// TIA Portal project "OP-TQ-01" (V13) (continued)
REGION Network 24: RESET ALARME DE SINAL ANALÓGICO
   RUNG wire#powerrail
      I_Contact( #Alarms.LL )
      I_Contact( #Alarms.L )
      I_Contact( #Alarms.H )
      I_Contact( #Alarms.HH )
      Contact( #RESET )
      wire#w1
      R_Coil( #AnalogInputAlarm )
   END_RUNG
   RUNG wire#powerrail
      Contact( #UnableAlarms )
   END_RUNG wire#w1
   RUNG wire#powerrail
      Contact( #Maint )
   END_RUNG wire#w1
   // the same network as SCL:
   IF (NOT #Alarms.LL AND NOT #Alarms.L AND NOT #Alarms.H AND NOT #Alarms.HH AND #RESET) OR #UnableAlarms OR #Maint THEN
       #AnalogInputAlarm := FALSE;
   END_IF;
END_REGION

REGION Network 25: 0 - STATUS OK
   RUNG wire#powerrail
      I_Contact( #AnalogInputFault )
      I_Contact( #AnalogInputAlarm )
      Contact( #Maint )
      { S7_GenerateENO := "TRUE" } Move(in := 0, out1 => #Status)
   END_RUNG
   // the same network as SCL:
   IF NOT #AnalogInputFault AND NOT #AnalogInputAlarm AND #Maint THEN #Status := 0; END_IF;
END_REGION

REGION Network 26: 1 - STATUS FALHA - UNDER FLOW
   RUNG wire#powerrail
      Contact( #Alarms.UDF )
      Contact( #Maint )
      { S7_GenerateENO := "TRUE" } Move(in := 1, out1 => #Status)
   END_RUNG
   // the same network as SCL:
   IF #Alarms.UDF AND #Maint THEN #Status := 1; END_IF;
END_REGION

REGION Network 27: 2 - STATUS FALHA - UNDER RANGE
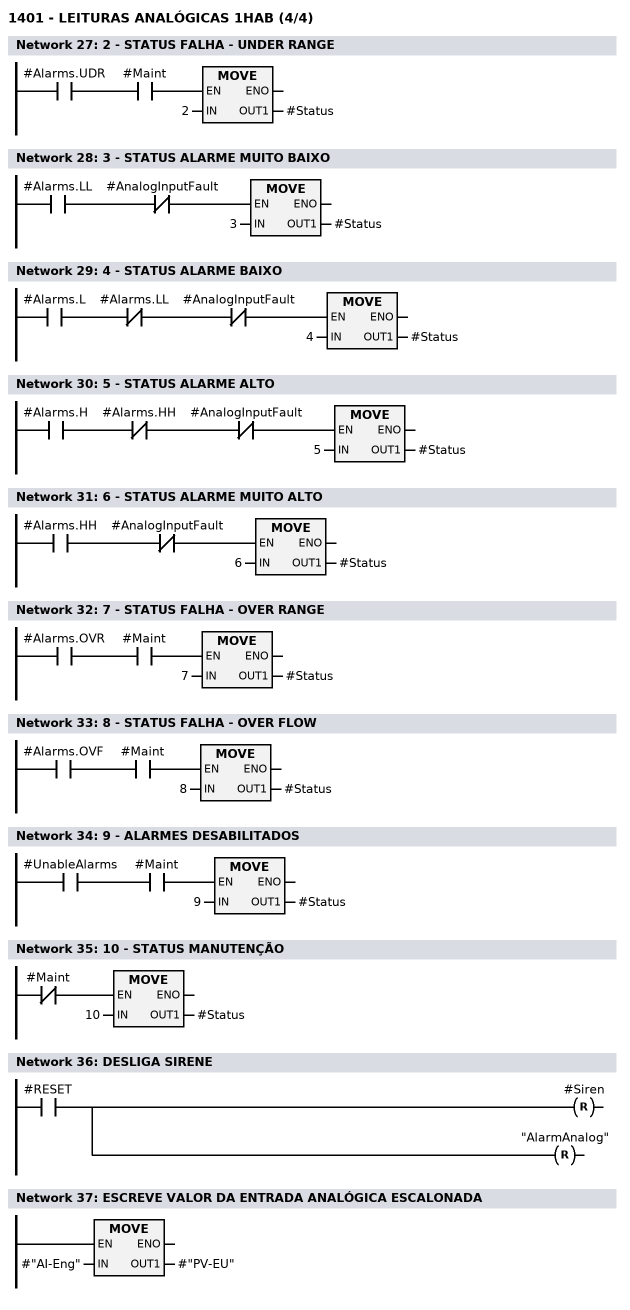
   RUNG wire#powerrail
      Contact( #Alarms.UDR )
      Contact( #Maint )
      { S7_GenerateENO := "TRUE" } Move(in := 2, out1 => #Status)
   END_RUNG
   // the same network as SCL:
   IF #Alarms.UDR AND #Maint THEN #Status := 2; END_IF;
END_REGION

REGION Network 28: 3 - STATUS ALARME MUITO BAIXO
   RUNG wire#powerrail
      Contact( #Alarms.LL )
      I_Contact( #AnalogInputFault )
      { S7_GenerateENO := "TRUE" } Move(in := 3, out1 => #Status)
   END_RUNG
   // the same network as SCL:
   IF #Alarms.LL AND NOT #AnalogInputFault THEN #Status := 3; END_IF;
END_REGION

REGION Network 29: 4 - STATUS ALARME BAIXO
   RUNG wire#powerrail
      Contact( #Alarms.L )
      I_Contact( #Alarms.LL )
      I_Contact( #AnalogInputFault )
      { S7_GenerateENO := "TRUE" } Move(in := 4, out1 => #Status)
   END_RUNG
   // the same network as SCL:
   IF #Alarms.L AND NOT #Alarms.LL AND NOT #AnalogInputFault THEN #Status := 4; END_IF;
END_REGION

REGION Network 30: 5 - STATUS ALARME ALTO
   RUNG wire#powerrail
      Contact( #Alarms.H )
      I_Contact( #Alarms.HH )
      I_Contact( #AnalogInputFault )
      { S7_GenerateENO := "TRUE" } Move(in := 5, out1 => #Status)
   END_RUNG
   // the same network as SCL:
   IF #Alarms.H AND NOT #Alarms.HH AND NOT #AnalogInputFault THEN #Status := 5; END_IF;
END_REGION

REGION Network 31: 6 - STATUS ALARME MUITO ALTO
   RUNG wire#powerrail
      Contact( #Alarms.HH )
      I_Contact( #AnalogInputFault )
      { S7_GenerateENO := "TRUE" } Move(in := 6, out1 => #Status)
   END_RUNG
   // the same network as SCL:
   IF #Alarms.HH AND NOT #AnalogInputFault THEN #Status := 6; END_IF;
END_REGION

REGION Network 32: 7 - STATUS FALHA - OVER RANGE
   RUNG wire#powerrail
      Contact( #Alarms.OVR )
      Contact( #Maint )
      { S7_GenerateENO := "TRUE" } Move(in := 7, out1 => #Status)
   END_RUNG
   // the same network as SCL:
   IF #Alarms.OVR AND #Maint THEN #Status := 7; END_IF;
END_REGION

REGION Network 33: 8 - STATUS FALHA - OVER FLOW
   RUNG wire#powerrail
      Contact( #Alarms.OVF )
      Contact( #Maint )
      { S7_GenerateENO := "TRUE" } Move(in := 8, out1 => #Status)
   END_RUNG
   // the same network as SCL:
   IF #Alarms.OVF AND #Maint THEN #Status := 8; END_IF;
END_REGION

REGION Network 34: 9 - ALARMES DESABILITADOS
   RUNG wire#powerrail
      Contact( #UnableAlarms )
      Contact( #Maint )
      { S7_GenerateENO := "TRUE" } Move(in := 9, out1 => #Status)
   END_RUNG
   // the same network as SCL:
   IF #UnableAlarms AND #Maint THEN #Status := 9; END_IF;
END_REGION

REGION Network 35: 10 - STATUS MANUTENÇÃO
   RUNG wire#powerrail
      I_Contact( #Maint )
      { S7_GenerateENO := "TRUE" } Move(in := 10, out1 => #Status)
   END_RUNG
   // the same network as SCL:
   IF NOT #Maint THEN #Status := 10; END_IF;
END_REGION

REGION Network 36: DESLIGA SIRENE
   RUNG wire#powerrail
      Contact( #RESET )
      wire#w1
      R_Coil( #Siren )
   END_RUNG
   RUNG wire#w1
      R_Coil( "AlarmAnalog" )
   END_RUNG
   // the same network as SCL:
   IF #RESET THEN
       #Siren := FALSE;
       "AlarmAnalog" := FALSE;
   END_IF;
END_REGION

REGION Network 37: ESCREVE VALOR DA ENTRADA ANALÓGICA ESCALONADA
   RUNG wire#powerrail
      { S7_GenerateENO := "TRUE" } Move(in := #"AI-Eng", out1 => #"PV-EU")
   END_RUNG
   // the same network as SCL:
   #"PV-EU" := #"AI-Eng";
END_REGION
END_FUNCTION_BLOCK

FUNCTION "1500 - SP-TT" : Void   // FC1500, LAD
{ S7_Optimized_Access := 'FALSE' }
VERSION : 0.1
   VAR_TEMP   // added for the SCL form of the ladder/FBD networks
      _w1 : Bool;
   END_VAR
BEGIN

REGION Network 1: VERIFICA TEMPERATURA MAX MAIOR QUE MIN
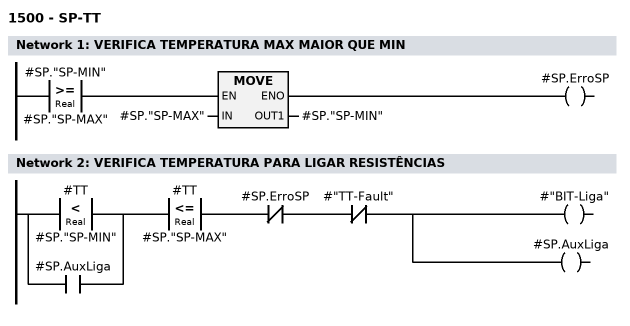
   RUNG wire#powerrail
      { S7_Templates := "SrcType := Real" } GE_Contact(in1 := #SP."SP-MIN", in2 := #SP."SP-MAX")
      { S7_GenerateENO := "TRUE" } Move(in := #SP."SP-MAX", out1 => #SP."SP-MIN")
      Coil( #SP.ErroSP )
   END_RUNG
   // the same network as SCL:
   // ENO of a box is taken as its EN; it also drops when the box reports an error
   #_w1 := #SP."SP-MIN" >= #SP."SP-MAX";
   IF #_w1 THEN #SP."SP-MIN" := #SP."SP-MAX"; END_IF;
   #SP.ErroSP := #_w1;
END_REGION

REGION Network 2: VERIFICA TEMPERATURA PARA LIGAR RESISTÊNCIAS
   RUNG wire#powerrail
      { S7_Templates := "SrcType := Real" } LT_Contact(in1 := #TT, in2 := #SP."SP-MIN")
      wire#w1
      { S7_Templates := "SrcType := Real" } LE_Contact(in1 := #TT, in2 := #SP."SP-MAX")
      I_Contact( #SP.ErroSP )
      I_Contact( #"TT-Fault" )
      wire#w2
      Coil( #"BIT-Liga" )
   END_RUNG
   RUNG wire#powerrail
      Contact( #SP.AuxLiga )
   END_RUNG wire#w1
   RUNG wire#w2
      Coil( #SP.AuxLiga )
   END_RUNG
   // the same network as SCL:
   #"BIT-Liga" := ((#TT < #SP."SP-MIN") OR #SP.AuxLiga) AND (#TT <= #SP."SP-MAX") AND NOT #SP.ErroSP AND NOT #"TT-Fault";
   #SP.AuxLiga := #"BIT-Liga";
END_REGION
END_FUNCTION

(* ===== HMI "HMI_RT_1" =====
connection "HMI_Connection_1": ETHERNET, S7_1200_OMS

HMI tags "Default tag table"
   "REC_ALM" : Bool = PLC "REC_ALM", 1 s
   "TT-006-R01A_AlarmsSts" : Alm-Bits, 1 s
   "TT-007-R01B_AlarmsSts" : Alm-Bits, 1 s
   "TT-008-R01C_AlarmsSts" : Alm-Bits, 1 s
   "TT-009-R01D_AlarmsSts" : Alm-Bits, 1 s
   "TT-010-R01E_AlarmsSts" : Alm-Bits, 1 s
   "TT-011-R01F_AlarmsSts" : Alm-Bits, 1 s
   "LT-009_AlarmsSts" : Alm-Bits, 1 s
   "LT-008_AlarmsSts" : Alm-Bits, 1 s

HMI tags "TT-006-R01A"
   "TT-006-R01A_UnableAlarms" : Bool, 1 s
   "TT-006-R01A_EngMax" : Real, 1 s
   "TT-006-R01A_EngMin" : Real, 1 s
   "TT-006-R01A_SP-HH" : Real, 1 s
   "TT-006-R01A_SP-H" : Real, 1 s
   "TT-006-R01A_SP-L" : Real, 1 s
   "TT-006-R01A_SP-LL" : Real, 1 s
   "TT-006-R01A_DelayHH" : Time, 1 s
   "TT-006-R01A_DelayH" : Time, 1 s
   "TT-006-R01A_DelayL" : Time, 1 s
   "TT-006-R01A_DelayLL" : Time, 1 s
   "TT-006-R01A_Siren" : Bool, 1 s
   "TT-006-R01A_SupRESET" : Bool, 1 s
   "TT-006-R01A_maint" : Bool, 1 s
   "TT-006-R01A_AlarmsEnable" : Alm-Bits, 1 s
   "TT-006-R01A_Alarms" : Alm-Bits, 1 s
   "TT-006-R01A_AI-Eng" : Real, 1 s
   "TT-006-R01A_Status" : Int, 1 s
   "TT-006-R01A_AnalogInput" : Int, 1 s

HMI tags "TT-007-R01B"
   "TT-007-R01B_UnableAlarms" : Bool, 1 s
   "TT-007-R01B_EngMax" : Real, 1 s
   "TT-007-R01B_EngMin" : Real, 1 s
   "TT-007-R01B_SP-HH" : Real, 1 s
   "TT-007-R01B_SP-H" : Real, 1 s
   "TT-007-R01B_SP-L" : Real, 1 s
   "TT-007-R01B_SP-LL" : Real, 1 s
   "TT-007-R01B_DelayHH" : Time, 1 s
   "TT-007-R01B_DelayH" : Time, 1 s
   "TT-007-R01B_DelayL" : Time, 1 s
   "TT-007-R01B_DelayLL" : Time, 1 s
   "TT-007-R01B_Siren" : Bool, 1 s
   "TT-007-R01B_SupRESET" : Bool, 1 s
   "TT-007-R01B_maint" : Bool, 1 s
   "TT-007-R01B_AlarmsEnable" : Alm-Bits, 1 s
   "TT-007-R01B_Alarms" : Alm-Bits, 1 s
   "TT-007-R01B_AI-Eng" : Real, 1 s
   "TT-007-R01B_Status" : Int, 1 s
   "TT-007-R01B_AnalogInput" : Int, 1 s

HMI tags "TT-008-R01C"
   "TT-008-R01C_UnableAlarms" : Bool, 1 s
   "TT-008-R01C_EngMax" : Real, 1 s
   "TT-008-R01C_EngMin" : Real, 1 s
   "TT-008-R01C_SP-HH" : Real, 1 s
   "TT-008-R01C_SP-H" : Real, 1 s
   "TT-008-R01C_SP-L" : Real, 1 s
   "TT-008-R01C_SP-LL" : Real, 1 s
   "TT-008-R01C_DelayHH" : Time, 1 s
   "TT-008-R01C_DelayH" : Time, 1 s
   "TT-008-R01C_DelayL" : Time, 1 s
   "TT-008-R01C_DelayLL" : Time, 1 s
   "TT-008-R01C_Siren" : Bool, 1 s
   "TT-008-R01C_SupRESET" : Bool, 1 s
   "TT-008-R01C_maint" : Bool, 1 s
   "TT-008-R01C_AlarmsEnable" : Alm-Bits, 1 s
   "TT-008-R01C_Alarms" : Alm-Bits, 1 s
   "TT-008-R01C_AI-Eng" : Real, 1 s
   "TT-008-R01C_Status" : Int, 1 s
   "TT-008-R01C_AnalogInput" : Int, 1 s

HMI tags "TT-009-R01D"
   "TT-009-R01D_UnableAlarms" : Bool, 1 s
   "TT-009-R01D_EngMax" : Real, 1 s
   "TT-009-R01D_EngMin" : Real, 1 s
   "TT-009-R01D_SP-HH" : Real, 1 s
   "TT-009-R01D_SP-H" : Real, 1 s
   "TT-009-R01D_SP-L" : Real, 1 s
   "TT-009-R01D_SP-LL" : Real, 1 s
   "TT-009-R01D_DelayHH" : Time, 1 s
   "TT-009-R01D_DelayH" : Time, 1 s
   "TT-009-R01D_DelayL" : Time, 1 s
   "TT-009-R01D_DelayLL" : Time, 1 s
   "TT-009-R01D_Siren" : Bool, 1 s
   "TT-009-R01D_SupRESET" : Bool, 1 s
   "TT-009-R01D_maint" : Bool, 1 s
   "TT-009-R01D_AlarmsEnable" : Alm-Bits, 1 s
   "TT-009-R01D_Alarms" : Alm-Bits, 1 s
   "TT-009-R01D_AI-Eng" : Real, 1 s
   "TT-009-R01D_Status" : Int, 1 s
   "TT-009-R01D_AnalogInput" : Int, 1 s

HMI tags "TT-010-R01E"
   "TT-010-R01E_UnableAlarms" : Bool, 1 s
   "TT-010-R01E_EngMax" : Real, 1 s
   "TT-010-R01E_EngMin" : Real, 1 s
   "TT-010-R01E_SP-HH" : Real, 1 s
   "TT-010-R01E_SP-H" : Real, 1 s
   "TT-010-R01E_SP-L" : Real, 1 s
   "TT-010-R01E_SP-LL" : Real, 1 s
   "TT-010-R01E_DelayHH" : Time, 1 s
   "TT-010-R01E_DelayH" : Time, 1 s
   "TT-010-R01E_DelayL" : Time, 1 s
   "TT-010-R01E_DelayLL" : Time, 1 s
   "TT-010-R01E_Siren" : Bool, 1 s
   "TT-010-R01E_SupRESET" : Bool, 1 s
   "TT-010-R01E_maint" : Bool, 1 s
   "TT-010-R01E_AlarmsEnable" : Alm-Bits, 1 s
   "TT-010-R01E_Alarms" : Alm-Bits, 1 s
   "TT-010-R01E_AI-Eng" : Real, 1 s
   "TT-010-R01E_Status" : Int, 1 s
   "TT-010-R01E_AnalogInput" : Int, 1 s

HMI tags "TT-011-R01F"
   "TT-011-R01F_UnableAlarms" : Bool, 1 s
   "TT-011-R01F_EngMax" : Real, 1 s
   "TT-011-R01F_EngMin" : Real, 1 s
   "TT-011-R01F_SP-HH" : Real, 1 s
   "TT-011-R01F_SP-H" : Real, 1 s
   "TT-011-R01F_SP-L" : Real, 1 s
   "TT-011-R01F_SP-LL" : Real, 1 s
   "TT-011-R01F_DelayHH" : Time, 1 s
   "TT-011-R01F_DelayH" : Time, 1 s
   "TT-011-R01F_DelayL" : Time, 1 s
   "TT-011-R01F_DelayLL" : Time, 1 s
   "TT-011-R01F_Siren" : Bool, 1 s
   "TT-011-R01F_SupRESET" : Bool, 1 s
   "TT-011-R01F_maint" : Bool, 1 s
   "TT-011-R01F_AlarmsEnable" : Alm-Bits, 1 s
   "TT-011-R01F_Alarms" : Alm-Bits, 1 s
   "TT-011-R01F_AI-Eng" : Real, 1 s
   "TT-011-R01F_Status" : Int, 1 s
   "TT-011-R01F_AnalogInput" : Int, 1 s

HMI tags "LT-009"
   "LT-009_UnableAlarms" : Bool, 1 s
   "LT-009_EngMax" : Real, 1 s
   "LT-009_EngMin" : Real, 1 s
   "LT-009_SP-HH" : Real, 1 s
   "LT-009_SP-H" : Real, 1 s
   "LT-009_SP-L" : Real, 1 s
   "LT-009_SP-LL" : Real, 1 s
   "LT-009_DelayHH" : Time, 1 s
   "LT-009_DelayH" : Time, 1 s
   "LT-009_DelayL" : Time, 1 s
   "LT-009_DelayLL" : Time, 1 s
   "LT-009_Siren" : Bool, 1 s
   "LT-009_SupRESET" : Bool, 1 s
   "LT-009_maint" : Bool, 1 s
   "LT-009_AlarmsEnable" : Alm-Bits, 1 s
   "LT-009_Alarms" : Alm-Bits, 1 s
   "LT-009_AI-Eng" : Real, 1 s
   "LT-009_Status" : Int, 1 s
   "LT-009_AnalogInput" : Int, 1 s

HMI tags "LT-008"
   "LT-008_UnableAlarms" : Bool, 1 s
   "LT-008_EngMax" : Real, 1 s
   "LT-008_EngMin" : Real, 1 s
   "LT-008_SP-HH" : Real, 1 s
   "LT-008_SP-H" : Real, 1 s
   "LT-008_SP-L" : Real, 1 s
   "LT-008_SP-LL" : Real, 1 s
   "LT-008_DelayHH" : Time, 1 s
   "LT-008_DelayH" : Time, 1 s
   "LT-008_DelayL" : Time, 1 s
   "LT-008_DelayLL" : Time, 1 s
   "LT-008_Siren" : Bool, 1 s
   "LT-008_SupRESET" : Bool, 1 s
   "LT-008_maint" : Bool, 1 s
   "LT-008_AlarmsEnable" : Alm-Bits, 1 s
   "LT-008_Alarms" : Alm-Bits, 1 s
   "LT-008_AI-Eng" : Real, 1 s
   "LT-008_Status" : Int, 1 s
   "LT-008_AnalogInput" : Int, 1 s

HMI tags "R01A-R01F"
   "R01A-R01F_BIT-Auto" : Bool, 1 s
   "R01A-R01F_Status" : Int, 1 s
   "R01A-R01F_OpTimeMinutes" : DInt, 1 s
   "R01A-R01F_OpTimeHours" : DInt, 1 s
   "R01A-R01F_SupRESET" : Bool, 1 s
   "R01A-R01F_Alm_Thermic" : Bool, 1 s
   "R01A-R01F_Alm_Interlock" : Bool, 1 s
   "R01A-R01F_Alm_FaultON" : Bool, 1 s
   "R01A-R01F_Alm_FaultOFF" : Bool, 1 s
   "R01A-R01F_FirstFault" : Int, 1 s
   "R01A-R01F_Command" : Int, 1 s
   "R01A-R01F_AutoMan" : Int, 1 s
   "R01A-R01F_StartCounter" : DInt, 1 s
   "SP-TT_TT-006-R01A" : SP-Temperaturas, 1 s
   "SP-TT_TT-007-R01B" : SP-Temperaturas, 1 s
   "SP-TT_TT-008-R01C" : SP-Temperaturas, 1 s
   "SP-TT_TT-009-R01D" : SP-Temperaturas, 1 s
   "SP-TT_TT-010-R01E" : SP-Temperaturas, 1 s
   "SP-TT_TT-011-R01F" : SP-Temperaturas, 1 s
   "R01A-R01F_SeletoraLR" : Bool, 1 s

HMI tags "ALARMES"
   "ALM_LSLL-004" : Bool, 1 s
   "ALM_TSH-004" : Bool, 1 s
   "ALM_FaltaDeFase" : Bool, 1 s
   "ALARMES-1" : UInt, 1 s
   "TT-006-R01A_Alarmes" : UInt, 1 s
   "TT-007-R01B_Alarmes" : UInt, 1 s
   "TT-008-R01C_Alarmes" : UInt, 1 s
   "TT-009-R01D_Alarmes" : UInt, 1 s
   "TT-010-R01E_Alarmes" : UInt, 1 s
   "TT-011-R01F_Alarmes" : UInt, 1 s
   "LT-009_Alarmes" : UInt, 1 s
   "LT-008_Alarmes" : UInt, 1 s

discrete alarms
   1: '', class Errors, trigger "ALARMES-1" bit 8
   2: '', class Errors, trigger "ALARMES-1" bit 9
   3: '', class Errors, trigger "ALARMES-1" bit 10
   4: '', class Errors, trigger "TT-006-R01A_Alarmes" bit 12
   5: '', class Errors, trigger "TT-006-R01A_Alarmes" bit 13
   6: '', class Errors, trigger "TT-006-R01A_Alarmes" bit 14
   7: '', class Errors, trigger "TT-006-R01A_Alarmes" bit 15
   8: '', class Errors, trigger "TT-007-R01B_Alarmes" bit 14
   9: '', class Errors, trigger "TT-007-R01B_Alarmes" bit 15
   10: '', class Errors, trigger "TT-007-R01B_Alarmes" bit 12
   11: '', class Errors, trigger "TT-007-R01B_Alarmes" bit 13
   12: '', class Errors, trigger "TT-008-R01C_Alarmes" bit 14
   13: '', class Errors, trigger "TT-008-R01C_Alarmes" bit 15
   14: '', class Errors, trigger "TT-008-R01C_Alarmes" bit 12
   15: '', class Errors, trigger "TT-008-R01C_Alarmes" bit 13
   16: '', class Errors, trigger "TT-009-R01D_Alarmes" bit 14
   17: '', class Errors, trigger "TT-009-R01D_Alarmes" bit 15
   18: '', class Errors, trigger "TT-009-R01D_Alarmes" bit 12
   19: '', class Errors, trigger "TT-009-R01D_Alarmes" bit 13
   20: '', class Errors, trigger "TT-010-R01E_Alarmes" bit 14
   21: '', class Errors, trigger "TT-010-R01E_Alarmes" bit 15
   22: '', class Errors, trigger "TT-010-R01E_Alarmes" bit 12
   23: '', class Errors, trigger "TT-010-R01E_Alarmes" bit 13
   24: '', class Errors, trigger "TT-011-R01F_Alarmes" bit 14
   25: '', class Errors, trigger "TT-011-R01F_Alarmes" bit 15
   26: '', class Errors, trigger "TT-011-R01F_Alarmes" bit 12
   27: '', class Errors, trigger "TT-011-R01F_Alarmes" bit 13
   28: '', class Errors, trigger "LT-009_Alarmes" bit 14
   29: '', class Errors, trigger "LT-009_Alarmes" bit 15
   30: '', class Errors, trigger "LT-009_Alarmes" bit 12
   31: '', class Errors, trigger "LT-009_Alarmes" bit 13
   32: '', class Errors, trigger "LT-008_Alarmes" bit 14
   33: '', class Errors, trigger "LT-008_Alarmes" bit 15
   34: '', class Errors, trigger "LT-008_Alarmes" bit 12
   35: '', class Errors, trigger "LT-008_Alarmes" bit 13

text list "ESTADO": 0 ''; 1 ''; 2 ''; 3 ''; 4 ''

text list "LR": 0 ''; 1 ''

text list "AM": 0 ''; 1 ''

screen "0000 - Apresentação" 480x272, template "Template_1"
   Button "Button_1" at 20,155 size 100x55
   TextField "HmiScreenItemData" at 0,55 size 480x85
   Button "Button_3" at 135,155 size 100x55
   Button "Button_4" at 250,155 size 100x55
   Button "Button_2" at 365,155 size 100x55
   Button "Button_5" at 20,210 size 100x55
   Button "Button_6" at 135,210 size 100x55

screen "1201 - TQ-OP-01" 480x272, template "Template_1"
   ScreenModuleView "EA-Painel-V_1" at 355,125 size 85x45
   ScreenModuleView "EA-Painel_1" at 10,55 size 170x26
   ScreenModuleView "EA-Painel_2" at 10,85 size 170x26
   ScreenModuleView "EA-Painel_3" at 10,115 size 170x26
   ScreenModuleView "EA-Painel_4" at 10,145 size 170x26
   ScreenModuleView "EA-Painel_5" at 10,175 size 170x26
   ScreenModuleView "EA-Painel_6" at 10,205 size 170x26
   TextField "HmiScreenItemData_4" at 215,130 size 15x15
   TextField "HmiScreenItemData_5" at 215,130 size 15x15
   TextField "HmiScreenItemData" at 75,5 size 225x30
   Bar "Bar_1" at 445,70 size 20x155
   TextField "HmiScreenItemData_8" at 290,55 size 95x25
   TextField "HmiScreenItemData_9" at 235,205 size 75x20
   TextField "HmiScreenItemData_1" at 235,175 size 75x20
   TextField "HmiScreenItemData_2" at 215,145 size 75x15
   Button "Button_3" at 265,240 size 65x32
   Button "Button_4" at 380,240 size 65x32
   Button "Button_1" at 295,95 size 40x30
   Button "Button_2" at 295,125 size 40x30
   GraphicView "Graphic view_1" at 275,105 size 15x15
   GraphicView "Graphic view_2" at 275,105 size 15x15
   TextField "HmiScreenItemData_10" at 275,130 size 15x15
   TextField "HmiScreenItemData_11" at 275,130 size 15x15
   SymbolicIOField "Symbolic I/O field_2" at 215,90 size 75x15

screen "1202 - BBC-OP-02" 480x272, template "Template_1"
   ScreenModuleView "EA-Painel-V_1" at 255,125 size 85x45
   Bar "Bar_1" at 345,70 size 20x155
   TextField "HmiScreenItemData_8" at 190,55 size 95x25
   TextField "HmiScreenItemData_9" at 135,205 size 75x20
   TextField "HmiScreenItemData_1" at 135,90 size 75x20
   TextField "HmiScreenItemData_2" at 135,115 size 75x20
   TextField "HmiScreenItemData_3" at 135,180 size 75x20

screen "System screens" 480x272, template "Template_1"
   TextField "HmiScreenItemData" at 48,93 size 384x22
   Button "HmiScreenItemData_1" at 1,1 size 157x36
   Button "HmiScreenItemData_2" at 159,1 size 157x36
   Button "HmiScreenItemData_3" at 317,1 size 157x36
   Button "HmiScreenItemData_4" at 1,38 size 157x36
   Button "HmiScreenItemData_5" at 159,38 size 157x36
   Button "HmiScreenItemData_6" at 317,38 size 157x36

screen "SIMATIC PLC system diagnostics" 480x272, template "Template_1"
   SysDiagControl "HmiScreenItemData" at 1,38 size 476x168
   Button "HmiScreenItemData_1" at 1,1 size 157x36

screen "Project information" 480x272, template "Template_1"
   TextField "HmiScreenItemData" at 4,39 size 184x20
   TextField "HmiScreenItemData_1" at 192,39 size 284x20
   TextField "HmiScreenItemData_2" at 4,60 size 184x20
   TextField "HmiScreenItemData_3" at 192,60 size 284x20
   TextField "HmiScreenItemData_4" at 4,81 size 184x20
   TextField "HmiScreenItemData_5" at 192,81 size 284x20
   TextField "HmiScreenItemData_6" at 4,102 size 184x20
   TextField "HmiScreenItemData_7" at 192,102 size 284x20
   Button "HmiScreenItemData_8" at 1,1 size 157x36

screen "User administration" 480x272, template "Template_1"
   UserView "HmiScreenItemData" at 1,38 size 476x168
   Button "HmiScreenItemData_1" at 1,1 size 157x36

screen "System information" 480x272, template "Template_1"
   TextField "HmiScreenItemData" at 4,39 size 184x20
   TextField "HmiScreenItemData_1" at 192,39 size 284x20
   TextField "HmiScreenItemData_2" at 4,60 size 184x20
   TextField "HmiScreenItemData_3" at 4,81 size 184x20
   TextField "HmiScreenItemData_4" at 192,81 size 284x20
   TextField "HmiScreenItemData_5" at 4,102 size 184x20
   TextField "HmiScreenItemData_6" at 192,102 size 284x20
   Button "HmiScreenItemData_7" at 192,60 size 284x20
   Button "HmiScreenItemData_8" at 1,1 size 157x36

screen "Different jobs" 480x272, template "Template_1"
   Button "HmiScreenItemData" at 1,38 size 157x36
   Button "HmiScreenItemData_1" at 1,75 size 157x36
   Button "HmiScreenItemData_2" at 1,112 size 157x36
   Button "HmiScreenItemData_3" at 1,149 size 157x36
   Button "HmiScreenItemData_4" at 159,38 size 157x36
   Button "HmiScreenItemData_5" at 159,75 size 157x36
   Button "HmiScreenItemData_6" at 1,1 size 157x36

screen "1301 - ALARMES" 480x272, template "Template_1"
   AlarmView "Alarm view_1" at 0,0 size 480x272

screen "1413 - TT-008-R01C" 480x272, template "Template_1"
   TextField "HmiScreenItemData" at 75,5 size 225x30
   ScreenModuleView "Ent-Analog_1" at 5,45 size 465x220

screen "1412 - TT-007-R01B" 480x272, template "Template_1"
   ScreenModuleView "Ent-Analog_1" at 5,45 size 465x220
   TextField "HmiScreenItemData" at 75,5 size 225x30

screen "1415 - TT-010-R01E" 480x272, template "Template_1"
   TextField "HmiScreenItemData" at 75,5 size 225x30
   ScreenModuleView "Ent-Analog_1" at 5,45 size 465x220

screen "1414 - TT-009-R01D" 480x272, template "Template_1"
   TextField "HmiScreenItemData" at 75,5 size 225x30
   ScreenModuleView "Ent-Analog_1" at 5,45 size 465x220

screen "1416 - TT-011-R01F" 480x272, template "Template_1"
   TextField "HmiScreenItemData" at 75,5 size 225x30
   ScreenModuleView "Ent-Analog_1" at 5,45 size 465x220

screen "1417 - LT-009" 480x272, template "Template_1"
   TextField "HmiScreenItemData" at 75,5 size 225x30
   ScreenModuleView "Ent-Analog_1" at 5,45 size 465x220

screen "1418 - LT-008" 480x272, template "Template_1"
   TextField "HmiScreenItemData" at 75,5 size 225x30
   ScreenModuleView "Ent-Analog_1" at 5,45 size 465x220

screen "1101 - Resistências" 480x272, template "Template_1"
   Button "Button_1" at 35,220 size 65x52
   TextField "HmiScreenItemData" at 75,5 size 225x30
   Button "Button_2" at 150,220 size 65x52
   SymbolicIOField "Symbolic I/O field_1" at 170,45 size 120x20
   TextField "HmiScreenItemData_1" at 305,45 size 170x20
   TextField "AlarmeUDF" at 325,65 size 150x20
   TextField "AlarmeUDF_1" at 325,105 size 150x20
   TextField "AlarmeUDF_2" at 325,85 size 150x20
   TextField "AlarmeUDF_3" at 325,125 size 150x20
   TextField "HmiScreenItemData_2" at 175,130 size 110x20
   TextField "HmiScreenItemData_3" at 220,145 size 15x20
   TextField "HmiScreenItemData_6" at 255,145 size 30x20
   IOField "I/O field_2" at 175,145 size 45x20
   IOField "I/O field_1" at 235,145 size 20x20
   TextField "HmiScreenItemData_7" at 170,165 size 120x30
   IOField "I/O field_3" at 170,190 size 120x20
   Button "Button_3" at 260,220 size 65x52
   TextField "HmiScreenItemData_8" at 310,150 size 160x20
   TextField "AlarmeUDF_4" at 355,170 size 70x15
   TextField "AlarmeUDF_5" at 355,185 size 70x15
   TextField "AlarmeUDF_6" at 355,200 size 70x15
   TextField "AlarmeUDF_7" at 355,215 size 70x15
   TextField "AlarmeUDF_8" at 355,230 size 70x15
   TextField "AlarmeUDF_9" at 355,245 size 70x15
   TextField "HmiScreenItemData_9" at 5,60 size 150x20
   TextField "AlarmeUDF_10" at 5,80 size 75x15
   TextField "AlarmeUDF_11" at 80,80 size 75x15
   TextField "AlarmeUDF_12" at 5,95 size 75x15
   TextField "AlarmeUDF_13" at 80,95 size 75x15
   TextField "AlarmeUDF_14" at 5,110 size 75x15
   TextField "AlarmeUDF_15" at 80,110 size 75x15
   TextField "AlarmeUDF_16" at 5,125 size 150x15
   TextField "AlarmeUDF_17" at 5,155 size 150x15
   TextField "AlarmeUDF_18" at 5,170 size 150x15
   TextField "AlarmeUDF_19" at 5,140 size 150x15
   GraphicView "Graphic view_3" at 270,65 size 20x20
   GraphicView "Graphic view_4" at 270,65 size 20x20
   TextField "HmiScreenItemData_4" at 170,105 size 20x20
   TextField "HmiScreenItemData_5" at 170,105 size 20x20
   TextField "HmiScreenItemData_10" at 270,105 size 20x20
   TextField "HmiScreenItemData_11" at 285,150 size 20x20

screen "1411 - TT-006-R01A" 480x272, template "Template_1"
   ScreenModuleView "Ent-Analog_1" at 5,45 size 465x220
   TextField "HmiScreenItemData" at 75,5 size 225x30

screen "1501 - SP" 480x272, template "Template_1"
   TextField "HmiScreenItemData" at 75,5 size 225x30
   ScreenModuleView "RESIST-SP_1" at 20,55 size 200x60
   ScreenModuleView "RESIST-SP_7" at 260,55 size 200x60
   ScreenModuleView "RESIST-SP_2" at 20,120 size 200x60
   ScreenModuleView "RESIST-SP_3" at 260,120 size 200x60
   ScreenModuleView "RESIST-SP_4" at 20,185 size 200x60
   ScreenModuleView "RESIST-SP_5" at 260,185 size 200x60

screen "1401 - ANALOG-MANUTENÇÃO" 480x272, template "Template_1"
   Button "Button_1" at 20,155 size 100x55
   TextField "HmiScreenItemData" at 0,45 size 480x85
   Button "Button_3" at 135,155 size 100x55
   Button "Button_4" at 250,155 size 100x55
   Button "Button_2" at 365,155 size 100x55
   Button "Button_5" at 20,210 size 100x55
   Button "Button_6" at 135,210 size 100x55
   Button "Button_7" at 250,210 size 100x55
   Button "Button_8" at 365,210 size 100x55

Template "Template_1" 480x272
   GraphicView "Template_Graphic view_1" at 300,0 size 180x40
   DateTimeField "Template_Date/time field_1" at 0,0 size 80x20
   DateTimeField "Template_Date/time field_2" at 0,20 size 80x20
*)

(* ===== HMI "HMI_RT_1" =====

ScreenModuleEditorView "EA-Painel-V" 640x480
   IOField "Indicador-Analogico" at 10,35 size 85x25
   TextField "TAG-Txt" at 10,15 size 85x20
*)

(* ===== HMI "HMI_RT_1" =====

ScreenModuleEditorView "EA-Painel" 640x480
   IOField "Indicador-Analogico" at 100,10 size 80x25
   TextField "TAG-Txt" at 10,10 size 90x25
*)

(* ===== HMI "HMI_RT_1" =====

ScreenModuleEditorView "Ent-Analog" 640x480
   TextField "F1-Txt" at 280,25 size 140x40
   TextField "F2-Txt" at 280,70 size 40x40
   TextField "Desab-Txt" at 307,70 size 113x40
   Button "F2-DesabAlarmes" at 280,70 size 140x40
   Button "F1-Manut" at 280,25 size 140x40
   IOField "Indicador-Analogico" at 145,10 size 110x35
   GraphicView "Alert-OFF-H" at 395,140 size 25x25
   GraphicView "Alert-OFF-L" at 395,165 size 25x25
   GraphicView "Alert-ON-H" at 395,140 size 25x25
   GraphicView "Alert-ON-L" at 395,165 size 25x25
   GraphicView "AlarmeOFF-HH" at 395,115 size 25x25
   GraphicView "AlarmeOFF-LL" at 395,190 size 25x25
   GraphicView "AlarmeON-HH" at 395,115 size 25x25
   GraphicView "AlarmeON-LL" at 395,190 size 25x25
   GraphicView "SireneOff" at 425,60 size 50x50
   GraphicView "AlarmeOff" at 385,75 size 30x30
   TextField "TAG-Txt" at 10,10 size 135x35
   IOField "EA-Bruta" at 153,85 size 70x25
   TextField "EA-Bruta-Txt" at 43,85 size 110x25
   IOField "SP-HH" at 310,115 size 80x25
   IOField "SP-H" at 310,140 size 80x25
   IOField "SP-L" at 310,165 size 80x25
   IOField "SP-LL" at 310,190 size 80x25
   GraphicView "AlarmeOn" at 385,75 size 30x30
   TextField "AlarmHabilitado-HH" at 280,115 size 30x25
   TextField "AlarmHabilitado-H" at 280,140 size 30x25
   TextField "AlarmHabilitado-L" at 280,165 size 30x25
   TextField "AlarmHabilitado-LL" at 280,190 size 30x25
   TextField "Alarmes-Lista-Txt" at 35,110 size 195x25
   TextField "AlarmeUDF" at 65,135 size 160x20
   TextField "AlarmeUDR" at 65,160 size 160x20
   TextField "AlarmeOVR" at 65,185 size 160x20
   TextField "AlarmeOVF" at 65,210 size 160x20
   GraphicView "Manut-Icone" at 390,30 size 25x30
   TextField "EngMin-Txt" at 10,50 size 50x25
   IOField "EngMin" at 60,50 size 70x25
   TextField "EngMax-Txt" at 135,50 size 50x25
   IOField "EngMax" at 185,50 size 70x25
   IOField "Tempo-HH" at 425,115 size 50x25
   IOField "Tempo-H" at 425,140 size 50x25
   IOField "Tempo-L" at 425,165 size 50x25
   IOField "Tempo-LL" at 425,190 size 50x25
   GraphicView "SireneOn" at 425,60 size 50x50
   TextField "F4-Txt" at 425,25 size 50x35
   Button "F4-Reset" at 425,25 size 50x85
   GraphicView "UDF-OFF" at 35,130 size 25x25
   GraphicView "UDF-ON" at 35,130 size 25x25
   GraphicView "UDR-OFF" at 35,155 size 25x25
   GraphicView "UDR-ON" at 35,155 size 25x25
   GraphicView "OVR-OFF" at 35,180 size 25x25
   GraphicView "OVR-ON" at 35,180 size 25x25
   GraphicView "OVF-OFF" at 35,205 size 25x25
   GraphicView "OVF-ON" at 35,205 size 25x25
   Button "DesabUDF" at 35,130 size 25x25
   Button "DesabUDR" at 35,155 size 25x25
   Button "DesabOVR" at 35,180 size 25x25
   Button "DesabOFV" at 35,205 size 25x25
*)

(* ===== HMI "HMI_RT_1" =====

ScreenModuleEditorView "RESIST-SP" 640x480
   TextField "TXT-MIN" at 10,55 size 120x20
   IOField "SP-MAX" at 130,35 size 80x20
   IOField "Indicador-Analogico" at 120,15 size 90x20
   TextField "TAG-Txt" at 10,15 size 110x20
   TextField "TXT-MAX" at 10,35 size 120x20
   IOField "SP-MIN" at 130,55 size 80x20
*)

(* ===== HMI "HMI_RT_1" =====

ScreenModuleEditorView "Ent-Analog" 640x480
   GraphicView "Alert-OFF-H" at 395,140 size 25x25
   GraphicView "Alert-OFF-L" at 395,165 size 25x25
   GraphicView "AlarmeOFF-HH" at 395,115 size 25x25
   GraphicView "AlarmeOFF-LL" at 395,190 size 25x25
   GraphicView "Alert-ON-H" at 395,140 size 25x25
   GraphicView "Alert-ON-L" at 395,165 size 25x25
   GraphicView "AlarmeON-HH" at 395,115 size 25x25
   GraphicView "AlarmeON-LL" at 395,190 size 25x25
   TextField "F1-Txt" at 280,25 size 140x40
   TextField "F2-Txt" at 280,70 size 40x40
   TextField "Desab-Txt" at 307,70 size 113x40
   Button "F2-DesabAlarmes" at 280,70 size 140x40
   Button "F1-Manut" at 280,25 size 140x40
   IOField "Indicador-Analogico" at 145,10 size 110x35
   GraphicView "SireneOff" at 425,60 size 50x50
   GraphicView "AlarmeOff" at 385,75 size 30x30
   TextField "TAG-Txt" at 10,10 size 135x35
   IOField "EA-Bruta" at 153,85 size 70x25
   TextField "EA-Bruta-Txt" at 43,85 size 110x25
   IOField "SP-HH" at 310,115 size 80x25
   IOField "SP-H" at 310,140 size 80x25
   IOField "SP-L" at 310,165 size 80x25
   IOField "SP-LL" at 310,190 size 80x25
   GraphicView "AlarmeOn" at 385,75 size 30x30
   TextField "AlarmHabilitado-HH" at 280,115 size 30x25
   TextField "AlarmHabilitado-H" at 280,140 size 30x25
   TextField "AlarmHabilitado-L" at 280,165 size 30x25
   TextField "AlarmHabilitado-LL" at 280,190 size 30x25
   TextField "Alarmes-Lista-Txt" at 35,110 size 195x25
   TextField "AlarmeUDF" at 65,135 size 160x20
   TextField "AlarmeUDR" at 65,160 size 160x20
   TextField "AlarmeOVR" at 65,185 size 160x20
   TextField "AlarmeOVF" at 65,210 size 160x20
   GraphicView "Manut-Icone" at 390,30 size 25x30
   TextField "EngMin-Txt" at 10,50 size 50x25
   IOField "EngMin" at 60,50 size 70x25
   TextField "EngMax-Txt" at 135,50 size 50x25
   IOField "EngMax" at 185,50 size 70x25
   IOField "Tempo-HH" at 425,115 size 50x25
   IOField "Tempo-H" at 425,140 size 50x25
   IOField "Tempo-L" at 425,165 size 50x25
   IOField "Tempo-LL" at 425,190 size 50x25
   GraphicView "SireneOn" at 425,60 size 50x50
   TextField "F4-Txt" at 425,25 size 50x35
   Button "F4-Reset" at 425,25 size 50x85
   GraphicView "UDF-OFF" at 35,130 size 25x25
   GraphicView "UDF-ON" at 35,130 size 25x25
   GraphicView "UDR-OFF" at 35,155 size 25x25
   GraphicView "UDR-ON" at 35,155 size 25x25
   GraphicView "OVR-OFF" at 35,180 size 25x25
   GraphicView "OVR-ON" at 35,180 size 25x25
   GraphicView "OVF-OFF" at 35,205 size 25x25
   GraphicView "OVF-ON" at 35,205 size 25x25
   Button "DesabUDF" at 35,130 size 25x25
   Button "DesabUDR" at 35,155 size 25x25
   Button "DesabOVR" at 35,180 size 25x25
   Button "DesabOFV" at 35,205 size 25x25
*)

(* ===== HMI "HMI_RT_1" =====

ScreenModuleEditorView "Ent-Analog" 640x480
   GraphicView "Alert-OFF-H" at 395,140 size 25x25
   GraphicView "Alert-OFF-L" at 395,165 size 25x25
   GraphicView "AlarmeOFF-HH" at 395,115 size 25x25
   GraphicView "AlarmeOFF-LL" at 395,190 size 25x25
   GraphicView "Alert-ON-H" at 395,140 size 25x25
   GraphicView "Alert-ON-L" at 395,165 size 25x25
   GraphicView "AlarmeON-HH" at 395,115 size 25x25
   GraphicView "AlarmeON-LL" at 395,190 size 25x25
   TextField "F1-Txt" at 280,25 size 140x40
   TextField "F2-Txt" at 280,70 size 40x40
   TextField "Desab-Txt" at 307,70 size 113x40
   Button "F2-DesabAlarmes" at 280,70 size 140x40
   Button "F1-Manut" at 280,25 size 140x40
   IOField "Indicador-Analogico" at 145,10 size 110x35
   GraphicView "SireneOff" at 425,60 size 50x50
   GraphicView "AlarmeOff" at 385,75 size 30x30
   TextField "TAG-Txt" at 10,10 size 135x35
   IOField "EA-Bruta" at 153,85 size 70x25
   TextField "EA-Bruta-Txt" at 43,85 size 110x25
   IOField "SP-HH" at 310,115 size 80x25
   IOField "SP-H" at 310,140 size 80x25
   IOField "SP-L" at 310,165 size 80x25
   IOField "SP-LL" at 310,190 size 80x25
   GraphicView "AlarmeOn" at 385,75 size 30x30
   TextField "AlarmHabilitado-HH" at 280,115 size 30x25
   TextField "AlarmHabilitado-H" at 280,140 size 30x25
   TextField "AlarmHabilitado-L" at 280,165 size 30x25
   TextField "AlarmHabilitado-LL" at 280,190 size 30x25
   TextField "Alarmes-Lista-Txt" at 35,110 size 195x25
   TextField "AlarmeUDF" at 65,135 size 160x20
   TextField "AlarmeUDR" at 65,160 size 160x20
   TextField "AlarmeOVR" at 65,185 size 160x20
   TextField "AlarmeOVF" at 65,210 size 160x20
   GraphicView "Manut-Icone" at 390,30 size 25x30
   TextField "EngMin-Txt" at 10,50 size 50x25
   IOField "EngMin" at 60,50 size 70x25
   TextField "EngMax-Txt" at 135,50 size 50x25
   IOField "EngMax" at 185,50 size 70x25
   IOField "Tempo-HH" at 425,115 size 50x25
   IOField "Tempo-H" at 425,140 size 50x25
   IOField "Tempo-L" at 425,165 size 50x25
   IOField "Tempo-LL" at 425,190 size 50x25
   GraphicView "SireneOn" at 425,60 size 50x50
   TextField "F4-Txt" at 425,25 size 50x35
   Button "F4-Reset" at 425,25 size 50x85
   GraphicView "UDF-OFF" at 35,130 size 25x25
   GraphicView "UDF-ON" at 35,130 size 25x25
   GraphicView "UDR-OFF" at 35,155 size 25x25
   GraphicView "UDR-ON" at 35,155 size 25x25
   GraphicView "OVR-OFF" at 35,180 size 25x25
   GraphicView "OVR-ON" at 35,180 size 25x25
   GraphicView "OVF-OFF" at 35,205 size 25x25
   GraphicView "OVF-ON" at 35,205 size 25x25
   Button "DesabUDF" at 35,130 size 25x25
   Button "DesabUDR" at 35,155 size 25x25
   Button "DesabOVR" at 35,180 size 25x25
   Button "DesabOFV" at 35,205 size 25x25
*)